   "Carrier_55_FaultLight_LH" AT %I3118.1 : Bool;   // FAULT LIGHT LH
   "Carrier_55_RunLight_LH" AT %I3118.2 : Bool;   // RUN LIGHT LH
   "Carrier_55_FaultLight_RH" AT %I3118.3 : Bool;   // FAULT LIGHT RH
   "Carrier_55_RunLight_RH" AT %I3118.4 : Bool;   // RUN LIGHT RH
   "Carrier_55_SpareOutput(5_5)" AT %I3118.5 : Bool;   // SPARE OUTPUT
   "Carrier_55_SpareOutput(5_6)" AT %I3118.6 : Bool;   // SPARE OUTPUT
   "Carrier_55_SpareOutput(5_7)" AT %I3118.7 : Bool;   // SPARE OUTPUT
   "Carrier_55_ActualSpeed" AT %IW3120 : Word;   // ACTUAL SPEED
   "Carrier_55_CarrierDriveAlarm" AT %IW3122 : Word;   // CARRIER DRIVE ALARM
   "Carrier_55_CarrierDriveWarning" AT %IW3124 : Word;   // CARRIER DRIVE WARNING
   "Carrier_56_Status" AT %IW3150 : Word;   // CARRIER STATUS WORD
   "Carrier_56_Status.0" AT %I3150.0 : Bool;   // HEARTBEAT
   "Carrier_56_Status.1" AT %I3150.1 : Bool;   // MANUAL
   "Carrier_56_Status.2" AT %I3150.2 : Bool;   // IN_AUTO
   "Carrier_56_Status.3" AT %I3150.3 : Bool;   // POSITIONING_COMPLETE
   "Carrier_56_Status.4" AT %I3150.4 : Bool;   // PRODUCTION HOLD
   "Carrier_56_Status.5" AT %I3150.5 : Bool;   // CARRIER MOVING FORWARD
   "Carrier_56_Status.6" AT %I3150.6 : Bool;   // CARRIER MOVING REVERSE
   "Carrier_56_Status.7" AT %I3150.7 : Bool;   // CARRIER FAULT
   "Carrier_56_Status.8" AT %I3151.0 : Bool;   // CRASH DETECT TRIPPED
   "Carrier_56_Status.9" AT %I3151.1 : Bool;
   "Carrier_56_Status.10" AT %I3151.2 : Bool;
   "Carrier_56_Status.11" AT %I3151.3 : Bool;
   "Carrier_56_Status.12" AT %I3151.4 : Bool;
   "Carrier_56_Status.13" AT %I3151.5 : Bool;
   "Carrier_56_Status.14" AT %I3151.6 : Bool;
   "Carrier_56_Status.15" AT %I3151.7 : Bool;
   "Carrier_56_SDCFaultCode" AT %IW3152 : Word;   // SDC FAULT CODE
   "Carrier_56_CarrierPosition" AT %ID3154 : DWord;   // CARRIER POSITION
   "Carrier_56_CarrierNumber" AT %IW3158 : Word;   // CARRIER NUMBER
   "Carrier_56_G120DControlWord" AT %IW3160 : Word;   // G120D_STW1_CONTROL
   "Carrier_56_G120DControlWord.0" AT %I3160.0 : Bool;   // Bit_00_ON
   "Carrier_56_G120DControlWord.1" AT %I3160.1 : Bool;   // Bit_01_AUS2_INH
   "Carrier_56_G120DControlWord.2" AT %I3160.2 : Bool;   // Bit_02_AUS3_STOP
   "Carrier_56_G120DControlWord.3" AT %I3160.3 : Bool;   // Bit_03_EN
   "Carrier_56_G120DControlWord.4" AT %I3160.4 : Bool;   // Bit_04_EN_RAMP
   "Carrier_56_G120DControlWord.5" AT %I3160.5 : Bool;   // Bit_05_START_RAMP
   "Carrier_56_G120DControlWord.6" AT %I3160.6 : Bool;   // Bit_06_SETPOINT
   "Carrier_56_G120DControlWord.7" AT %I3160.7 : Bool;   // Bit_07_RESET
   "Carrier_56_G120DControlWord.8" AT %I3161.0 : Bool;   // Bit_08_JOG_R
   "Carrier_56_G120DControlWord.9" AT %I3161.1 : Bool;   // Bit_09_JOG_L
   "Carrier_56_G120DControlWord.10" AT %I3161.2 : Bool;   // Bit_10_CONTR_PLC
   "Carrier_56_G120DControlWord.11" AT %I3161.3 : Bool;   // Bit_11_REVERSE
   "Carrier_56_G120DControlWord.12" AT %I3161.4 : Bool;   // Bit_12_BRAKE_RELEASE
   "Carrier_56_G120DControlWord.13" AT %I3161.5 : Bool;   // Bit_13_DDS
   "Carrier_56_G120DControlWord.14" AT %I3161.6 : Bool;   // Bit_14_DO0
   "Carrier_56_G120DControlWord.15" AT %I3161.7 : Bool;   // Bit_15_DO1
   "Carrier_56_G120DStatusWord" AT %IW3162 : Word;   // G120D_ZSW1_STATUS
   "Carrier_56_G120DStatusWord.0" AT %I3162.0 : Bool;   // Bit_00_READY_RUN
   "Carrier_56_G120DStatusWord.1" AT %I3162.1 : Bool;   // Bit_01_READY_ON
   "Carrier_56_G120DStatusWord.2" AT %I3162.2 : Bool;   // Bit_02_ENABLE
   "Carrier_56_G120DStatusWord.3" AT %I3162.3 : Bool;   // Bit_03_FAULT
   "Carrier_56_G120DStatusWord.4" AT %I3162.4 : Bool;   // Bit_04_OFF2
   "Carrier_56_G120DStatusWord.5" AT %I3162.5 : Bool;   // Bit_05_OFF3
   "Carrier_56_G120DStatusWord.6" AT %I3162.6 : Bool;   // Bit_06_LOCK_OUT
   "Carrier_56_G120DStatusWord.7" AT %I3162.7 : Bool;   // Bit_07_WARN
   "Carrier_56_G120DStatusWord.8" AT %I3163.0 : Bool;   // Bit_08_NO_DEVIATION
   "Carrier_56_G120DStatusWord.9" AT %I3163.1 : Bool;   // Bit_09_CONTR_PLC
   "Carrier_56_G120DStatusWord.10" AT %I3163.2 : Bool;   // Bit_10_F_MAX
   "Carrier_56_G120DStatusWord.11" AT %I3163.3 : Bool;   // Bit_11_LIMIT_REACHED
   "Carrier_56_G120DStatusWord.12" AT %I3163.4 : Bool;   // Bit_12_BRAKE_OPEN
   "Carrier_56_G120DStatusWord.13" AT %I3163.5 : Bool;   // Bit_13_NO_OVERTEMP
   "Carrier_56_G120DStatusWord.14" AT %I3163.6 : Bool;   // Bit_14_CW_CCW
   "Carrier_56_G120DStatusWord.15" AT %I3163.7 : Bool;   // Bit_15_OVERL
   "Carrier_56_Slot2_Input" AT %IW3164 : Word;   // SLOT 2 INPUT WORD
   "Carrier_56_CrashDetectSW" AT %I3164.0 : Bool;   // CRASH DETECT SW
   "Carrier_56_SpareSafetyInput(2_1)" AT %I3164.1 : Bool;   // SPARE SAFETY INPUT
   "Carrier_56_SpareSafetyInput(2_2)" AT %I3164.2 : Bool;   // SPARE SAFETY INPUT
   "Carrier_56_SpareSafetyInput(2_3)" AT %I3164.3 : Bool;   // SPARE SAFETY INPUT
   "Carrier_56_SpareSafetyInput(2_4)" AT %I3164.4 : Bool;   // SPARE SAFETY INPUT
   "Carrier_56_SpareSafetyInput(2_5)" AT %I3164.5 : Bool;   // SPARE SAFETY INPUT
   "Carrier_56_SpareSafetyInput(2_6)" AT %I3164.6 : Bool;   // SPARE SAFETY INPUT
   "Carrier_56_SpareSafetyInput(2_7)" AT %I3164.7 : Bool;   // SPARE SAFETY INPUT
   "Carrier_56_Slot3_SafetyOutput" AT %IW3165 : Word;   // SLOT 3 SAFETY OUTPUT WORD
   "Carrier_56_Crash_Detect_OK" AT %I3165.0 : Bool;   // CARRIER CRASH DETECT
   "Carrier_56_SpareSafetyOutput(3_1)" AT %I3165.1 : Bool;   // SPARE SAFETY OUTPUT
   "Carrier_56_SpareSafetyOutput(3_2)" AT %I3165.2 : Bool;   // SPARE SAFETY OUTPUT
   "Carrier_56_SpareSafetyOutput(3_3)" AT %I3165.3 : Bool;   // SPARE SAFETY OUTPUT
   "Carrier_56_SpareSafetyOutput(3_4)" AT %I3165.4 : Bool;   // SPARE SAFETY OUTPUT
   "Carrier_56_SpareSafetyOutput(3_5)" AT %I3165.5 : Bool;   // SPARE SAFETY OUTPUT
   "Carrier_56_SpareSafetyOutput(3_6)" AT %I3165.6 : Bool;   // SPARE SAFETY OUTPUT
   "Carrier_56_SpareSafetyOutput(3_7)" AT %I3165.7 : Bool;   // SPARE SAFETY OUTPUT
   "Carrier_56_Slot4_Input" AT %IW3166 : Word;   // SLOT 4 INPUT WORD
   "Carrier_56_480VPowerOn_MDCB1" AT %I3166.0 : Bool;   // 480 VAC POWER ON MDCB 1
   "Carrier_56_SpareInput(4_1)" AT %I3166.1 : Bool;   // SPARE INPUT
   "Carrier_56_SpareInput(4_2)" AT %I3166.2 : Bool;   // SPARE INPUT
   "Carrier_56_SitopSelectStatus" AT %I3166.3 : Bool;   // SITOP SELECT STATUS
   "Carrier_56_DCsupplyOnPSCB2" AT %I3166.4 : Bool;   // DC SUPPLY ON PSCB 2
   "Carrier_56_SpareInput(4_5)" AT %I3166.5 : Bool;   // SPARE INPUT
   "Carrier_56_SpareInput(4_6)" AT %I3166.6 : Bool;   // SPARE INPUT
   "Carrier_56_SpareInput(4_7)" AT %I3166.7 : Bool;   // SPARE INPUT
   "Carrier_56_PB1_ProdHoldLH" AT %I3167.0 : Bool;   // PB 1 PRODUCTION HOLD LH
   "Carrier_56_PB2_ResetLH" AT %I3167.1 : Bool;   // PB 2 RESET LH
   "Carrier_56_PB3_ProdHoldRH" AT %I3167.2 : Bool;   // PB 3 PRODUCTION HOLD RH
   "Carrier_56_PB4_ResetRH" AT %I3167.3 : Bool;   // PB 4 RESET RH
   "Carrier_56_SpareInput(4_14)" AT %I3167.4 : Bool;   // SPARE INPUT
   "Carrier_56_SpareInput(4_15)" AT %I3167.5 : Bool;   // SPARE INPUT
   "Carrier_56_SpareInput(4_16)" AT %I3167.6 : Bool;   // SPARE INPUT
   "Carrier_56_SpareInput(4_17)" AT %I3167.7 : Bool;   // SPARE INPUT
   "Carrier_56_Slot5_Output" AT %IW3168 : Word;   // SLOT 5 OUTPUT WORD
   "Carrier_56_IRD400_HMI_24VDC_ENABLE" AT %I3168.0 : Bool;   // IRD 400 PANEL HMI 24V DC POWER
   "Carrier_56_FaultLight_LH" AT %I3168.1 : Bool;   // FAULT LIGHT LH
   "Carrier_56_RunLight_LH" AT %I3168.2 : Bool;   // RUN LIGHT LH
   "Carrier_56_FaultLight_RH" AT %I3168.3 : Bool;   // FAULT LIGHT RH
   "Carrier_56_RunLight_RH" AT %I3168.4 : Bool;   // RUN LIGHT RH
   "Carrier_56_SpareOutput(5_5)" AT %I3168.5 : Bool;   // SPARE OUTPUT
   "Carrier_56_SpareOutput(5_6)" AT %I3168.6 : Bool;   // SPARE OUTPUT
   "Carrier_56_SpareOutput(5_7)" AT %I3168.7 : Bool;   // SPARE OUTPUT
   "Carrier_56_ActualSpeed" AT %IW3170 : Word;   // ACTUAL SPEED
   "Carrier_56_CarrierDriveAlarm" AT %IW3172 : Word;   // CARRIER DRIVE ALARM
   "Carrier_56_CarrierDriveWarning" AT %IW3174 : Word;   // CARRIER DRIVE WARNING
   "Carrier_57_Status" AT %IW3200 : Word;   // CARRIER STATUS WORD
   "Carrier_57_Status.0" AT %I3200.0 : Bool;   // HEARTBEAT
   "Carrier_57_Status.1" AT %I3200.1 : Bool;   // MANUAL
   "Carrier_57_Status.2" AT %I3200.2 : Bool;   // IN_AUTO
   "Carrier_57_Status.3" AT %I3200.3 : Bool;   // POSITIONING_COMPLETE
   "Carrier_57_Status.4" AT %I3200.4 : Bool;   // PRODUCTION HOLD
   "Carrier_57_Status.5" AT %I3200.5 : Bool;   // CARRIER MOVING FORWARD
   "Carrier_57_Status.6" AT %I3200.6 : Bool;   // CARRIER MOVING REVERSE
   "Carrier_57_Status.7" AT %I3200.7 : Bool;   // CARRIER FAULT
   "Carrier_57_Status.8" AT %I3201.0 : Bool;   // CRASH DETECT TRIPPED
   "Carrier_57_Status.9" AT %I3201.1 : Bool;
   "Carrier_57_Status.10" AT %I3201.2 : Bool;
   "Carrier_57_Status.11" AT %I3201.3 : Bool;
   "Carrier_57_Status.12" AT %I3201.4 : Bool;
   "Carrier_57_Status.13" AT %I3201.5 : Bool;
   "Carrier_57_Status.14" AT %I3201.6 : Bool;
   "Carrier_57_Status.15" AT %I3201.7 : Bool;
   "Carrier_57_SDCFaultCode" AT %IW3202 : Word;   // SDC FAULT CODE
   "Carrier_57_CarrierPosition" AT %ID3204 : DWord;   // CARRIER POSITION
   "Carrier_57_CarrierNumber" AT %IW3208 : Word;   // CARRIER NUMBER
   "Carrier_57_G120DControlWord" AT %IW3210 : Word;   // G120D_STW1_CONTROL
   "Carrier_57_G120DControlWord.0" AT %I3210.0 : Bool;   // Bit_00_ON
   "Carrier_57_G120DControlWord.1" AT %I3210.1 : Bool;   // Bit_01_AUS2_INH
   "Carrier_57_G120DControlWord.2" AT %I3210.2 : Bool;   // Bit_02_AUS3_STOP
   "Carrier_57_G120DControlWord.3" AT %I3210.3 : Bool;   // Bit_03_EN
   "Carrier_57_G120DControlWord.4" AT %I3210.4 : Bool;   // Bit_04_EN_RAMP
   "Carrier_57_G120DControlWord.5" AT %I3210.5 : Bool;   // Bit_05_START_RAMP
   "Carrier_57_G120DControlWord.6" AT %I3210.6 : Bool;   // Bit_06_SETPOINT
   "Carrier_57_G120DControlWord.7" AT %I3210.7 : Bool;   // Bit_07_RESET
   "Carrier_57_G120DControlWord.8" AT %I3211.0 : Bool;   // Bit_08_JOG_R
   "Carrier_57_G120DControlWord.9" AT %I3211.1 : Bool;   // Bit_09_JOG_L
   "Carrier_57_G120DControlWord.10" AT %I3211.2 : Bool;   // Bit_10_CONTR_PLC
   "Carrier_57_G120DControlWord.11" AT %I3211.3 : Bool;   // Bit_11_REVERSE
   "Carrier_57_G120DControlWord.12" AT %I3211.4 : Bool;   // Bit_12_BRAKE_RELEASE
   "Carrier_57_G120DControlWord.13" AT %I3211.5 : Bool;   // Bit_13_DDS
   "Carrier_57_G120DControlWord.14" AT %I3211.6 : Bool;   // Bit_14_DO0
   "Carrier_57_G120DControlWord.15" AT %I3211.7 : Bool;   // Bit_15_DO1
   "Carrier_57_G120DStatusWord" AT %IW3212 : Word;   // G120D_ZSW1_STATUS
   "Carrier_57_G120DStatusWord.0" AT %I3212.0 : Bool;   // Bit_00_READY_RUN
   "Carrier_57_G120DStatusWord.1" AT %I3212.1 : Bool;   // Bit_01_READY_ON
   "Carrier_57_G120DStatusWord.2" AT %I3212.2 : Bool;   // Bit_02_ENABLE
   "Carrier_57_G120DStatusWord.3" AT %I3212.3 : Bool;   // Bit_03_FAULT
   "Carrier_57_G120DStatusWord.4" AT %I3212.4 : Bool;   // Bit_04_OFF2
   "Carrier_57_G120DStatusWord.5" AT %I3212.5 : Bool;   // Bit_05_OFF3
   "Carrier_57_G120DStatusWord.6" AT %I3212.6 : Bool;   // Bit_06_LOCK_OUT
   "Carrier_57_G120DStatusWord.7" AT %I3212.7 : Bool;   // Bit_07_WARN
   "Carrier_57_G120DStatusWord.8" AT %I3213.0 : Bool;   // Bit_08_NO_DEVIATION
   "Carrier_57_G120DStatusWord.9" AT %I3213.1 : Bool;   // Bit_09_CONTR_PLC
   "Carrier_57_G120DStatusWord.10" AT %I3213.2 : Bool;   // Bit_10_F_MAX
   "Carrier_57_G120DStatusWord.11" AT %I3213.3 : Bool;   // Bit_11_LIMIT_REACHED
   "Carrier_57_G120DStatusWord.12" AT %I3213.4 : Bool;   // Bit_12_BRAKE_OPEN
   "Carrier_57_G120DStatusWord.13" AT %I3213.5 : Bool;   // Bit_13_NO_OVERTEMP
   "Carrier_57_G120DStatusWord.14" AT %I3213.6 : Bool;   // Bit_14_CW_CCW
   "Carrier_57_G120DStatusWord.15" AT %I3213.7 : Bool;   // Bit_15_OVERL
   "Carrier_57_Slot2_Input" AT %IW3214 : Word;   // SLOT 2 INPUT WORD
   "Carrier_57_CrashDetectSW" AT %I3214.0 : Bool;   // CRASH DETECT SW
   "Carrier_57_SpareSafetyInput(2_1)" AT %I3214.1 : Bool;   // SPARE SAFETY INPUT
   "Carrier_57_SpareSafetyInput(2_2)" AT %I3214.2 : Bool;   // SPARE SAFETY INPUT
   "Carrier_57_SpareSafetyInput(2_3)" AT %I3214.3 : Bool;   // SPARE SAFETY INPUT
   "Carrier_57_SpareSafetyInput(2_4)" AT %I3214.4 : Bool;   // SPARE SAFETY INPUT
   "Carrier_57_SpareSafetyInput(2_5)" AT %I3214.5 : Bool;   // SPARE SAFETY INPUT
   "Carrier_57_SpareSafetyInput(2_6)" AT %I3214.6 : Bool;   // SPARE SAFETY INPUT
   "Carrier_57_SpareSafetyInput(2_7)" AT %I3214.7 : Bool;   // SPARE SAFETY INPUT
   "Carrier_57_Slot3_SafetyOutput" AT %IW3215 : Word;   // SLOT 3 SAFETY OUTPUT WORD
   "Carrier_57_Crash_Detect_OK" AT %I3215.0 : Bool;   // CARRIER CRASH DETECT
   "Carrier_57_SpareSafetyOutput(3_1)" AT %I3215.1 : Bool;   // SPARE SAFETY OUTPUT
   "Carrier_57_SpareSafetyOutput(3_2)" AT %I3215.2 : Bool;   // SPARE SAFETY OUTPUT
   "Carrier_57_SpareSafetyOutput(3_3)" AT %I3215.3 : Bool;   // SPARE SAFETY OUTPUT
   "Carrier_57_SpareSafetyOutput(3_4)" AT %I3215.4 : Bool;   // SPARE SAFETY OUTPUT
   "Carrier_57_SpareSafetyOutput(3_5)" AT %I3215.5 : Bool;   // SPARE SAFETY OUTPUT
   "Carrier_57_SpareSafetyOutput(3_6)" AT %I3215.6 : Bool;   // SPARE SAFETY OUTPUT
   "Carrier_57_SpareSafetyOutput(3_7)" AT %I3215.7 : Bool;   // SPARE SAFETY OUTPUT
   "Carrier_57_Slot4_Input" AT %IW3216 : Word;   // SLOT 4 INPUT WORD
   "Carrier_57_480VPowerOn_MDCB1" AT %I3216.0 : Bool;   // 480 VAC POWER ON MDCB 1
   "Carrier_57_SpareInput(4_1)" AT %I3216.1 : Bool;   // SPARE INPUT
   "Carrier_57_SpareInput(4_2)" AT %I3216.2 : Bool;   // SPARE INPUT
   "Carrier_57_SitopSelectStatus" AT %I3216.3 : Bool;   // SITOP SELECT STATUS
   "Carrier_57_DCsupplyOnPSCB2" AT %I3216.4 : Bool;   // DC SUPPLY ON PSCB 2
   "Carrier_57_SpareInput(4_5)" AT %I3216.5 : Bool;   // SPARE INPUT
   "Carrier_57_SpareInput(4_6)" AT %I3216.6 : Bool;   // SPARE INPUT
   "Carrier_57_SpareInput(4_7)" AT %I3216.7 : Bool;   // SPARE INPUT
   "Carrier_57_PB1_ProdHoldLH" AT %I3217.0 : Bool;   // PB 1 PRODUCTION HOLD LH
   "Carrier_57_PB2_ResetLH" AT %I3217.1 : Bool;   // PB 2 RESET LH
   "Carrier_57_PB3_ProdHoldRH" AT %I3217.2 : Bool;   // PB 3 PRODUCTION HOLD RH
   "Carrier_57_PB4_ResetRH" AT %I3217.3 : Bool;   // PB 4 RESET RH
   "Carrier_57_SpareInput(4_14)" AT %I3217.4 : Bool;   // SPARE INPUT
   "Carrier_57_SpareInput(4_15)" AT %I3217.5 : Bool;   // SPARE INPUT
   "Carrier_57_SpareInput(4_16)" AT %I3217.6 : Bool;   // SPARE INPUT
   "Carrier_57_SpareInput(4_17)" AT %I3217.7 : Bool;   // SPARE INPUT
   "Carrier_57_Slot5_Output" AT %IW3218 : Word;   // SLOT 5 OUTPUT WORD
   "Carrier_57_IRD400_HMI_24VDC_ENABLE" AT %I3218.0 : Bool;   // IRD 400 PANEL HMI 24V DC POWER
   "Carrier_57_FaultLight_LH" AT %I3218.1 : Bool;   // FAULT LIGHT LH
   "Carrier_57_RunLight_LH" AT %I3218.2 : Bool;   // RUN LIGHT LH
   "Carrier_57_FaultLight_RH" AT %I3218.3 : Bool;   // FAULT LIGHT RH
   "Carrier_57_RunLight_RH" AT %I3218.4 : Bool;   // RUN LIGHT RH
   "Carrier_57_SpareOutput(5_5)" AT %I3218.5 : Bool;   // SPARE OUTPUT
   "Carrier_57_SpareOutput(5_6)" AT %I3218.6 : Bool;   // SPARE OUTPUT
   "Carrier_57_SpareOutput(5_7)" AT %I3218.7 : Bool;   // SPARE OUTPUT
   "Carrier_57_ActualSpeed" AT %IW3220 : Word;   // ACTUAL SPEED
   "Carrier_57_CarrierDriveAlarm" AT %IW3222 : Word;   // CARRIER DRIVE ALARM
   "Carrier_57_CarrierDriveWarning" AT %IW3224 : Word;   // CARRIER DRIVE WARNING
   "Carrier_58_Status" AT %IW3250 : Word;   // CARRIER STATUS WORD
   "Carrier_58_Status.0" AT %I3250.0 : Bool;   // HEARTBEAT
   "Carrier_58_Status.1" AT %I3250.1 : Bool;   // MANUAL
   "Carrier_58_Status.2" AT %I3250.2 : Bool;   // IN_AUTO
   "Carrier_58_Status.3" AT %I3250.3 : Bool;   // POSITIONING_COMPLETE
   "Carrier_58_Status.4" AT %I3250.4 : Bool;   // PRODUCTION HOLD
   "Carrier_58_Status.5" AT %I3250.5 : Bool;   // CARRIER MOVING FORWARD
   "Carrier_58_Status.6" AT %I3250.6 : Bool;   // CARRIER MOVING REVERSE
   "Carrier_58_Status.7" AT %I3250.7 : Bool;   // CARRIER FAULT
   "Carrier_58_Status.8" AT %I3251.0 : Bool;   // CRASH DETECT TRIPPED
   "Carrier_58_Status.9" AT %I3251.1 : Bool;
   "Carrier_58_Status.10" AT %I3251.2 : Bool;
   "Carrier_58_Status.11" AT %I3251.3 : Bool;
   "Carrier_58_Status.12" AT %I3251.4 : Bool;
   "Carrier_58_Status.13" AT %I3251.5 : Bool;
   "Carrier_58_Status.14" AT %I3251.6 : Bool;
   "Carrier_58_Status.15" AT %I3251.7 : Bool;
   "Carrier_58_SDCFaultCode" AT %IW3252 : Word;   // SDC FAULT CODE
   "Carrier_58_CarrierPosition" AT %ID3254 : DWord;   // CARRIER POSITION
   "Carrier_58_CarrierNumber" AT %IW3258 : Word;   // CARRIER NUMBER
   "Carrier_58_G120DControlWord" AT %IW3260 : Word;   // G120D_STW1_CONTROL
   "Carrier_58_G120DControlWord.0" AT %I3260.0 : Bool;   // Bit_00_ON
   "Carrier_58_G120DControlWord.1" AT %I3260.1 : Bool;   // Bit_01_AUS2_INH
   "Carrier_58_G120DControlWord.2" AT %I3260.2 : Bool;   // Bit_02_AUS3_STOP
   "Carrier_58_G120DControlWord.3" AT %I3260.3 : Bool;   // Bit_03_EN
   "Carrier_58_G120DControlWord.4" AT %I3260.4 : Bool;   // Bit_04_EN_RAMP
   "Carrier_58_G120DControlWord.5" AT %I3260.5 : Bool;   // Bit_05_START_RAMP
   "Carrier_58_G120DControlWord.6" AT %I3260.6 : Bool;   // Bit_06_SETPOINT
   "Carrier_58_G120DControlWord.7" AT %I3260.7 : Bool;   // Bit_07_RESET
   "Carrier_58_G120DControlWord.8" AT %I3261.0 : Bool;   // Bit_08_JOG_R
   "Carrier_58_G120DControlWord.9" AT %I3261.1 : Bool;   // Bit_09_JOG_L
   "Carrier_58_G120DControlWord.10" AT %I3261.2 : Bool;   // Bit_10_CONTR_PLC
   "Carrier_58_G120DControlWord.11" AT %I3261.3 : Bool;   // Bit_11_REVERSE
   "Carrier_58_G120DControlWord.12" AT %I3261.4 : Bool;   // Bit_12_BRAKE_RELEASE
   "Carrier_58_G120DControlWord.13" AT %I3261.5 : Bool;   // Bit_13_DDS
   "Carrier_58_G120DControlWord.14" AT %I3261.6 : Bool;   // Bit_14_DO0
   "Carrier_58_G120DControlWord.15" AT %I3261.7 : Bool;   // Bit_15_DO1
   "Carrier_58_G120DStatusWord" AT %IW3262 : Word;   // G120D_ZSW1_STATUS
   "Carrier_58_G120DStatusWord.0" AT %I3262.0 : Bool;   // Bit_00_READY_RUN
   "Carrier_58_G120DStatusWord.1" AT %I3262.1 : Bool;   // Bit_01_READY_ON
   "Carrier_58_G120DStatusWord.2" AT %I3262.2 : Bool;   // Bit_02_ENABLE
   "Carrier_58_G120DStatusWord.3" AT %I3262.3 : Bool;   // Bit_03_FAULT
   "Carrier_58_G120DStatusWord.4" AT %I3262.4 : Bool;   // Bit_04_OFF2
   "Carrier_58_G120DStatusWord.5" AT %I3262.5 : Bool;   // Bit_05_OFF3
   "Carrier_58_G120DStatusWord.6" AT %I3262.6 : Bool;   // Bit_06_LOCK_OUT
   "Carrier_58_G120DStatusWord.7" AT %I3262.7 : Bool;   // Bit_07_WARN
   "Carrier_58_G120DStatusWord.8" AT %I3263.0 : Bool;   // Bit_08_NO_DEVIATION
   "Carrier_58_G120DStatusWord.9" AT %I3263.1 : Bool;   // Bit_09_CONTR_PLC
   "Carrier_58_G120DStatusWord.10" AT %I3263.2 : Bool;   // Bit_10_F_MAX
   "Carrier_58_G120DStatusWord.11" AT %I3263.3 : Bool;   // Bit_11_LIMIT_REACHED
   "Carrier_58_G120DStatusWord.12" AT %I3263.4 : Bool;   // Bit_12_BRAKE_OPEN
   "Carrier_58_G120DStatusWord.13" AT %I3263.5 : Bool;   // Bit_13_NO_OVERTEMP
   "Carrier_58_G120DStatusWord.14" AT %I3263.6 : Bool;   // Bit_14_CW_CCW
   "Carrier_58_G120DStatusWord.15" AT %I3263.7 : Bool;   // Bit_15_OVERL
   "Carrier_58_Slot2_Input" AT %IW3264 : Word;   // SLOT 2 INPUT WORD
   "Carrier_58_CrashDetectSW" AT %I3264.0 : Bool;   // CRASH DETECT SW
   "Carrier_58_SpareSafetyInput(2_1)" AT %I3264.1 : Bool;   // SPARE SAFETY INPUT
   "Carrier_58_SpareSafetyInput(2_2)" AT %I3264.2 : Bool;   // SPARE SAFETY INPUT
   "Carrier_58_SpareSafetyInput(2_3)" AT %I3264.3 : Bool;   // SPARE SAFETY INPUT
   "Carrier_58_SpareSafetyInput(2_4)" AT %I3264.4 : Bool;   // SPARE SAFETY INPUT
   "Carrier_58_SpareSafetyInput(2_5)" AT %I3264.5 : Bool;   // SPARE SAFETY INPUT
   "Carrier_58_SpareSafetyInput(2_6)" AT %I3264.6 : Bool;   // SPARE SAFETY INPUT
   "Carrier_58_SpareSafetyInput(2_7)" AT %I3264.7 : Bool;   // SPARE SAFETY INPUT
   "Carrier_58_Slot3_SafetyOutput" AT %IW3265 : Word;   // SLOT 3 SAFETY OUTPUT WORD
   "Carrier_58_Crash_Detect_OK" AT %I3265.0 : Bool;   // CARRIER CRASH DETECT
   "Carrier_58_SpareSafetyOutput(3_1)" AT %I3265.1 : Bool;   // SPARE SAFETY OUTPUT
   "Carrier_58_SpareSafetyOutput(3_2)" AT %I3265.2 : Bool;   // SPARE SAFETY OUTPUT
   "Carrier_58_SpareSafetyOutput(3_3)" AT %I3265.3 : Bool;   // SPARE SAFETY OUTPUT
   "Carrier_58_SpareSafetyOutput(3_4)" AT %I3265.4 : Bool;   // SPARE SAFETY OUTPUT
   "Carrier_58_SpareSafetyOutput(3_5)" AT %I3265.5 : Bool;   // SPARE SAFETY OUTPUT
   "Carrier_58_SpareSafetyOutput(3_6)" AT %I3265.6 : Bool;   // SPARE SAFETY OUTPUT
   "Carrier_58_SpareSafetyOutput(3_7)" AT %I3265.7 : Bool;   // SPARE SAFETY OUTPUT
   "Carrier_58_Slot4_Input" AT %IW3266 : Word;   // SLOT 4 INPUT WORD
   "Carrier_58_480VPowerOn_MDCB1" AT %I3266.0 : Bool;   // 480 VAC POWER ON MDCB 1
   "Carrier_58_SpareInput(4_1)" AT %I3266.1 : Bool;   // SPARE INPUT
   "Carrier_58_SpareInput(4_2)" AT %I3266.2 : Bool;   // SPARE INPUT
   "Carrier_58_SitopSelectStatus" AT %I3266.3 : Bool;   // SITOP SELECT STATUS
   "Carrier_58_DCsupplyOnPSCB2" AT %I3266.4 : Bool;   // DC SUPPLY ON PSCB 2
   "Carrier_58_SpareInput(4_5)" AT %I3266.5 : Bool;   // SPARE INPUT
   "Carrier_58_SpareInput(4_6)" AT %I3266.6 : Bool;   // SPARE INPUT
   "Carrier_58_SpareInput(4_7)" AT %I3266.7 : Bool;   // SPARE INPUT
   "Carrier_58_PB1_ProdHoldLH" AT %I3267.0 : Bool;   // PB 1 PRODUCTION HOLD LH
   "Carrier_58_PB2_ResetLH" AT %I3267.1 : Bool;   // PB 2 RESET LH
   "Carrier_58_PB3_ProdHoldRH" AT %I3267.2 : Bool;   // PB 3 PRODUCTION HOLD RH
   "Carrier_58_PB4_ResetRH" AT %I3267.3 : Bool;   // PB 4 RESET RH
   "Carrier_58_SpareInput(4_14)" AT %I3267.4 : Bool;   // SPARE INPUT
   "Carrier_58_SpareInput(4_15)" AT %I3267.5 : Bool;   // SPARE INPUT
   "Carrier_58_SpareInput(4_16)" AT %I3267.6 : Bool;   // SPARE INPUT
   "Carrier_58_SpareInput(4_17)" AT %I3267.7 : Bool;   // SPARE INPUT
   "Carrier_58_Slot5_Output" AT %IW3268 : Word;   // SLOT 5 OUTPUT WORD
   "Carrier_58_IRD400_HMI_24VDC_ENABLE" AT %I3268.0 : Bool;   // IRD 400 PANEL HMI 24V DC POWER
   "Carrier_58_FaultLight_LH" AT %I3268.1 : Bool;   // FAULT LIGHT LH
   "Carrier_58_RunLight_LH" AT %I3268.2 : Bool;   // RUN LIGHT LH
   "Carrier_58_FaultLight_RH" AT %I3268.3 : Bool;   // FAULT LIGHT RH
   "Carrier_58_RunLight_RH" AT %I3268.4 : Bool;   // RUN LIGHT RH
   "Carrier_58_SpareOutput(5_5)" AT %I3268.5 : Bool;   // SPARE OUTPUT
   "Carrier_58_SpareOutput(5_6)" AT %I3268.6 : Bool;   // SPARE OUTPUT
   "Carrier_58_SpareOutput(5_7)" AT %I3268.7 : Bool;   // SPARE OUTPUT
   "Carrier_58_ActualSpeed" AT %IW3270 : Word;   // ACTUAL SPEED
   "Carrier_58_CarrierDriveAlarm" AT %IW3272 : Word;   // CARRIER DRIVE ALARM
   "Carrier_58_CarrierDriveWarning" AT %IW3274 : Word;   // CARRIER DRIVE WARNING
   "Carrier_59_Status" AT %IW3300 : Word;   // CARRIER STATUS WORD
   "Carrier_59_Status.0" AT %I3300.0 : Bool;   // HEARTBEAT
   "Carrier_59_Status.1" AT %I3300.1 : Bool;   // MANUAL
   "Carrier_59_Status.2" AT %I3300.2 : Bool;   // IN_AUTO
   "Carrier_59_Status.3" AT %I3300.3 : Bool;   // POSITIONING_COMPLETE
   "Carrier_59_Status.4" AT %I3300.4 : Bool;   // PRODUCTION HOLD
   "Carrier_59_Status.5" AT %I3300.5 : Bool;   // CARRIER MOVING FORWARD
   "Carrier_59_Status.6" AT %I3300.6 : Bool;   // CARRIER MOVING REVERSE
   "Carrier_59_Status.7" AT %I3300.7 : Bool;   // CARRIER FAULT
   "Carrier_59_Status.8" AT %I3301.0 : Bool;   // CRASH DETECT TRIPPED
   "Carrier_59_Status.9" AT %I3301.1 : Bool;
   "Carrier_59_Status.10" AT %I3301.2 : Bool;
   "Carrier_59_Status.11" AT %I3301.3 : Bool;
   "Carrier_59_Status.12" AT %I3301.4 : Bool;
   "Carrier_59_Status.13" AT %I3301.5 : Bool;
   "Carrier_59_Status.14" AT %I3301.6 : Bool;
   "Carrier_59_Status.15" AT %I3301.7 : Bool;
   "Carrier_59_SDCFaultCode" AT %IW3302 : Word;   // SDC FAULT CODE
   "Carrier_59_CarrierPosition" AT %ID3304 : DWord;   // CARRIER POSITION
   "Carrier_59_CarrierNumber" AT %IW3308 : Word;   // CARRIER NUMBER
   "Carrier_59_G120DControlWord" AT %IW3310 : Word;   // G120D_STW1_CONTROL
   "Carrier_59_G120DControlWord.0" AT %I3310.0 : Bool;   // Bit_00_ON
   "Carrier_59_G120DControlWord.1" AT %I3310.1 : Bool;   // Bit_01_AUS2_INH
   "Carrier_59_G120DControlWord.2" AT %I3310.2 : Bool;   // Bit_02_AUS3_STOP
   "Carrier_59_G120DControlWord.3" AT %I3310.3 : Bool;   // Bit_03_EN
   "Carrier_59_G120DControlWord.4" AT %I3310.4 : Bool;   // Bit_04_EN_RAMP
   "Carrier_59_G120DControlWord.5" AT %I3310.5 : Bool;   // Bit_05_START_RAMP
   "Carrier_59_G120DControlWord.6" AT %I3310.6 : Bool;   // Bit_06_SETPOINT
   "Carrier_59_G120DControlWord.7" AT %I3310.7 : Bool;   // Bit_07_RESET
   "Carrier_59_G120DControlWord.8" AT %I3311.0 : Bool;   // Bit_08_JOG_R
   "Carrier_59_G120DControlWord.9" AT %I3311.1 : Bool;   // Bit_09_JOG_L
   "Carrier_59_G120DControlWord.10" AT %I3311.2 : Bool;   // Bit_10_CONTR_PLC
   "Carrier_59_G120DControlWord.11" AT %I3311.3 : Bool;   // Bit_11_REVERSE
   "Carrier_59_G120DControlWord.12" AT %I3311.4 : Bool;   // Bit_12_BRAKE_RELEASE
   "Carrier_59_G120DControlWord.13" AT %I3311.5 : Bool;   // Bit_13_DDS
   "Carrier_59_G120DControlWord.14" AT %I3311.6 : Bool;   // Bit_14_DO0
   "Carrier_59_G120DControlWord.15" AT %I3311.7 : Bool;   // Bit_15_DO1
   "Carrier_59_G120DStatusWord" AT %IW3312 : Word;   // G120D_ZSW1_STATUS
   "Carrier_59_G120DStatusWord.0" AT %I3312.0 : Bool;   // Bit_00_READY_RUN
   "Carrier_59_G120DStatusWord.1" AT %I3312.1 : Bool;   // Bit_01_READY_ON
   "Carrier_59_G120DStatusWord.2" AT %I3312.2 : Bool;   // Bit_02_ENABLE
   "Carrier_59_G120DStatusWord.3" AT %I3312.3 : Bool;   // Bit_03_FAULT
   "Carrier_59_G120DStatusWord.4" AT %I3312.4 : Bool;   // Bit_04_OFF2
   "Carrier_59_G120DStatusWord.5" AT %I3312.5 : Bool;   // Bit_05_OFF3
   "Carrier_59_G120DStatusWord.6" AT %I3312.6 : Bool;   // Bit_06_LOCK_OUT
   "Carrier_59_G120DStatusWord.7" AT %I3312.7 : Bool;   // Bit_07_WARN
   "Carrier_59_G120DStatusWord.8" AT %I3313.0 : Bool;   // Bit_08_NO_DEVIATION
   "Carrier_59_G120DStatusWord.9" AT %I3313.1 : Bool;   // Bit_09_CONTR_PLC
   "Carrier_59_G120DStatusWord.10" AT %I3313.2 : Bool;   // Bit_10_F_MAX
   "Carrier_59_G120DStatusWord.11" AT %I3313.3 : Bool;   // Bit_11_LIMIT_REACHED
   "Carrier_59_G120DStatusWord.12" AT %I3313.4 : Bool;   // Bit_12_BRAKE_OPEN
   "Carrier_59_G120DStatusWord.13" AT %I3313.5 : Bool;   // Bit_13_NO_OVERTEMP
   "Carrier_59_G120DStatusWord.14" AT %I3313.6 : Bool;   // Bit_14_CW_CCW
   "Carrier_59_G120DStatusWord.15" AT %I3313.7 : Bool;   // Bit_15_OVERL
   "Carrier_59_Slot2_Input" AT %IW3314 : Word;   // SLOT 2 INPUT WORD
   "Carrier_59_CrashDetectSW" AT %I3314.0 : Bool;   // CRASH DETECT SW
   "Carrier_59_SpareSafetyInput(2_1)" AT %I3314.1 : Bool;   // SPARE SAFETY INPUT
   "Carrier_59_SpareSafetyInput(2_2)" AT %I3314.2 : Bool;   // SPARE SAFETY INPUT
   "Carrier_59_SpareSafetyInput(2_3)" AT %I3314.3 : Bool;   // SPARE SAFETY INPUT
   "Carrier_59_SpareSafetyInput(2_4)" AT %I3314.4 : Bool;   // SPARE SAFETY INPUT
   "Carrier_59_SpareSafetyInput(2_5)" AT %I3314.5 : Bool;   // SPARE SAFETY INPUT
   "Carrier_59_SpareSafetyInput(2_6)" AT %I3314.6 : Bool;   // SPARE SAFETY INPUT
   "Carrier_59_SpareSafetyInput(2_7)" AT %I3314.7 : Bool;   // SPARE SAFETY INPUT
   "Carrier_59_Slot3_SafetyOutput" AT %IW3315 : Word;   // SLOT 3 SAFETY OUTPUT WORD
   "Carrier_59_Crash_Detect_OK" AT %I3315.0 : Bool;   // CARRIER CRASH DETECT
   "Carrier_59_SpareSafetyOutput(3_1)" AT %I3315.1 : Bool;   // SPARE SAFETY OUTPUT
   "Carrier_59_SpareSafetyOutput(3_2)" AT %I3315.2 : Bool;   // SPARE SAFETY OUTPUT
   "Carrier_59_SpareSafetyOutput(3_3)" AT %I3315.3 : Bool;   // SPARE SAFETY OUTPUT
   "Carrier_59_SpareSafetyOutput(3_4)" AT %I3315.4 : Bool;   // SPARE SAFETY OUTPUT
   "Carrier_59_SpareSafetyOutput(3_5)" AT %I3315.5 : Bool;   // SPARE SAFETY OUTPUT
   "Carrier_59_SpareSafetyOutput(3_6)" AT %I3315.6 : Bool;   // SPARE SAFETY OUTPUT
   "Carrier_59_SpareSafetyOutput(3_7)" AT %I3315.7 : Bool;   // SPARE SAFETY OUTPUT
   "Carrier_59_Slot4_Input" AT %IW3316 : Word;   // SLOT 4 INPUT WORD
   "Carrier_59_480VPowerOn_MDCB1" AT %I3316.0 : Bool;   // 480 VAC POWER ON MDCB 1
   "Carrier_59_SpareInput(4_1)" AT %I3316.1 : Bool;   // SPARE INPUT
   "Carrier_59_SpareInput(4_2)" AT %I3316.2 : Bool;   // SPARE INPUT
   "Carrier_59_SitopSelectStatus" AT %I3316.3 : Bool;   // SITOP SELECT STATUS
   "Carrier_59_DCsupplyOnPSCB2" AT %I3316.4 : Bool;   // DC SUPPLY ON PSCB 2
   "Carrier_59_SpareInput(4_5)" AT %I3316.5 : Bool;   // SPARE INPUT
   "Carrier_59_SpareInput(4_6)" AT %I3316.6 : Bool;   // SPARE INPUT
   "Carrier_59_SpareInput(4_7)" AT %I3316.7 : Bool;   // SPARE INPUT
   "Carrier_59_PB1_ProdHoldLH" AT %I3317.0 : Bool;   // PB 1 PRODUCTION HOLD LH
   "Carrier_59_PB2_ResetLH" AT %I3317.1 : Bool;   // PB 2 RESET LH
   "Carrier_59_PB3_ProdHoldRH" AT %I3317.2 : Bool;   // PB 3 PRODUCTION HOLD RH
   "Carrier_59_PB4_ResetRH" AT %I3317.3 : Bool;   // PB 4 RESET RH
   "Carrier_59_SpareInput(4_14)" AT %I3317.4 : Bool;   // SPARE INPUT
   "Carrier_59_SpareInput(4_15)" AT %I3317.5 : Bool;   // SPARE INPUT
   "Carrier_59_SpareInput(4_16)" AT %I3317.6 : Bool;   // SPARE INPUT
   "Carrier_59_SpareInput(4_17)" AT %I3317.7 : Bool;   // SPARE INPUT
   "Carrier_59_Slot5_Output" AT %IW3318 : Word;   // SLOT 5 OUTPUT WORD
   "Carrier_59_IRD400_HMI_24VDC_ENABLE" AT %I3318.0 : Bool;   // IRD 400 PANEL HMI 24V DC POWER
   "Carrier_59_FaultLight_LH" AT %I3318.1 : Bool;   // FAULT LIGHT LH
   "Carrier_59_RunLight_LH" AT %I3318.2 : Bool;   // RUN LIGHT LH
   "Carrier_59_FaultLight_RH" AT %I3318.3 : Bool;   // FAULT LIGHT RH
   "Carrier_59_RunLight_RH" AT %I3318.4 : Bool;   // RUN LIGHT RH
   "Carrier_59_SpareOutput(5_5)" AT %I3318.5 : Bool;   // SPARE OUTPUT
   "Carrier_59_SpareOutput(5_6)" AT %I3318.6 : Bool;   // SPARE OUTPUT
   "Carrier_59_SpareOutput(5_7)" AT %I3318.7 : Bool;   // SPARE OUTPUT
   "Carrier_59_ActualSpeed" AT %IW3320 : Word;   // ACTUAL SPEED
   "Carrier_59_CarrierDriveAlarm" AT %IW3322 : Word;   // CARRIER DRIVE ALARM
   "Carrier_59_CarrierDriveWarning" AT %IW3324 : Word;   // CARRIER DRIVE WARNING
   "Carrier_60_Status" AT %IW3350 : Word;   // CARRIER STATUS WORD
   "Carrier_60_Status.0" AT %I3350.0 : Bool;   // HEARTBEAT
   "Carrier_60_Status.1" AT %I3350.1 : Bool;   // MANUAL
   "Carrier_60_Status.2" AT %I3350.2 : Bool;   // IN_AUTO
   "Carrier_60_Status.3" AT %I3350.3 : Bool;   // POSITIONING_COMPLETE
   "Carrier_60_Status.4" AT %I3350.4 : Bool;   // PRODUCTION HOLD
   "Carrier_60_Status.5" AT %I3350.5 : Bool;   // CARRIER MOVING FORWARD
   "Carrier_60_Status.6" AT %I3350.6 : Bool;   // CARRIER MOVING REVERSE
   "Carrier_60_Status.7" AT %I3350.7 : Bool;   // CARRIER FAULT
   "Carrier_60_Status.8" AT %I3351.0 : Bool;   // CRASH DETECT TRIPPED
   "Carrier_60_Status.9" AT %I3351.1 : Bool;
   "Carrier_60_Status.10" AT %I3351.2 : Bool;
   "Carrier_60_Status.11" AT %I3351.3 : Bool;
   "Carrier_60_Status.12" AT %I3351.4 : Bool;
   "Carrier_60_Status.13" AT %I3351.5 : Bool;
   "Carrier_60_Status.14" AT %I3351.6 : Bool;
   "Carrier_60_Status.15" AT %I3351.7 : Bool;
   "Carrier_60_SDCFaultCode" AT %IW3352 : Word;   // SDC FAULT CODE
   "Carrier_60_CarrierPosition" AT %ID3354 : DWord;   // CARRIER POSITION
   "Carrier_60_CarrierNumber" AT %IW3358 : Word;   // CARRIER NUMBER
   "Carrier_60_G120DControlWord" AT %IW3360 : Word;   // G120D_STW1_CONTROL
   "Carrier_60_G120DControlWord.0" AT %I3360.0 : Bool;   // Bit_00_ON
   "Carrier_60_G120DControlWord.1" AT %I3360.1 : Bool;   // Bit_01_AUS2_INH
   "Carrier_60_G120DControlWord.2" AT %I3360.2 : Bool;   // Bit_02_AUS3_STOP
   "Carrier_60_G120DControlWord.3" AT %I3360.3 : Bool;   // Bit_03_EN
   "Carrier_60_G120DControlWord.4" AT %I3360.4 : Bool;   // Bit_04_EN_RAMP
   "Carrier_60_G120DControlWord.5" AT %I3360.5 : Bool;   // Bit_05_START_RAMP
   "Carrier_60_G120DControlWord.6" AT %I3360.6 : Bool;   // Bit_06_SETPOINT
   "Carrier_60_G120DControlWord.7" AT %I3360.7 : Bool;   // Bit_07_RESET
   "Carrier_60_G120DControlWord.8" AT %I3361.0 : Bool;   // Bit_08_JOG_R
   "Carrier_60_G120DControlWord.9" AT %I3361.1 : Bool;   // Bit_09_JOG_L
   "Carrier_60_G120DControlWord.10" AT %I3361.2 : Bool;   // Bit_10_CONTR_PLC
   "Carrier_60_G120DControlWord.11" AT %I3361.3 : Bool;   // Bit_11_REVERSE
   "Carrier_60_G120DControlWord.12" AT %I3361.4 : Bool;   // Bit_12_BRAKE_RELEASE
   "Carrier_60_G120DControlWord.13" AT %I3361.5 : Bool;   // Bit_13_DDS
   "Carrier_60_G120DControlWord.14" AT %I3361.6 : Bool;   // Bit_14_DO0
   "Carrier_60_G120DControlWord.15" AT %I3361.7 : Bool;   // Bit_15_DO1
   "Carrier_60_G120DStatusWord" AT %IW3362 : Word;   // G120D_ZSW1_STATUS
   "Carrier_60_G120DStatusWord.0" AT %I3362.0 : Bool;   // Bit_00_READY_RUN
   "Carrier_60_G120DStatusWord.1" AT %I3362.1 : Bool;   // Bit_01_READY_ON
   "Carrier_60_G120DStatusWord.2" AT %I3362.2 : Bool;   // Bit_02_ENABLE
   "Carrier_60_G120DStatusWord.3" AT %I3362.3 : Bool;   // Bit_03_FAULT
   "Carrier_60_G120DStatusWord.4" AT %I3362.4 : Bool;   // Bit_04_OFF2
   "Carrier_60_G120DStatusWord.5" AT %I3362.5 : Bool;   // Bit_05_OFF3
   "Carrier_60_G120DStatusWord.6" AT %I3362.6 : Bool;   // Bit_06_LOCK_OUT
   "Carrier_60_G120DStatusWord.7" AT %I3362.7 : Bool;   // Bit_07_WARN
   "Carrier_60_G120DStatusWord.8" AT %I3363.0 : Bool;   // Bit_08_NO_DEVIATION
   "Carrier_60_G120DStatusWord.9" AT %I3363.1 : Bool;   // Bit_09_CONTR_PLC
   "Carrier_60_G120DStatusWord.10" AT %I3363.2 : Bool;   // Bit_10_F_MAX
   "Carrier_60_G120DStatusWord.11" AT %I3363.3 : Bool;   // Bit_11_LIMIT_REACHED